TYPE "typeMouldEditor_HMI"
VERSION : 0.1
   STRUCT
      sSelected : Struct   // Selected
         iTool : Int;   // Selected - tool
         sPS : Struct   // Selected - partial shot
            iPS : Int;
            arFlow : Array[0..6] of Real;
            arRatio : Array[0..6] of Real;
            arPressure : Array[0..6] of Real;
            RefComponent : Int;
            "2PoinMovement_Comp01" : Bool;
            "2PoinMovement_Comp02" : Bool;
            "2PoinMovement_Comp03" : Bool;
            "2PoinMovement_Comp04" : Bool;
            "2PoinMovement_Comp05" : Bool;
            "2PoinMovement_Comp06" : Bool;
         END_STRUCT;
         iCalculation : Int;   // Selected - calculation (0=Ftime; 1=flow; 2=weight)
      END_STRUCT;
      arShotSet : Array[0..8] of "UDT925_Shot";   // Shot settings
      uTools : "UDT930_Tool";   // Tool settings
      sCalculatedValues : Struct   // Calculated values
         arTotalFlow : Array[0..8] of Real;   // Calculated values - total flow
      END_STRUCT;
      sStatusBits : Struct   // StatusBits
         xValueChanged : Bool;   // Value changed
         xSafeChanges : Bool;   // Safe changes
         xDiscardChanges : Bool;   // Discard changes
         xDeleteProgram : Bool;   // Delete program
         xFaultDeleteProgram : Bool;   // Fault - delete program
         xProgLoadName : Bool;   // program load name
         xProgLoadNameAckn : Bool;   // program load name - acknowledge
         xFaultValuesnotvalid : Bool;   // values are not valid - flow or shot time wrong
         xPartShotAmount_increase : Bool;   // Partial shot amount - increase
         xPartShotAmount_decrease : Bool;   // Partial shot amount - decrease
      END_STRUCT;
      sColumn : Struct   // Column in HMI
         iShotTime : Int;   // Column - shot time
         iTotalFlow : Int;   // Column - total flow
         iTotalWeight : Int;   // Column - total weight
      END_STRUCT;
      sRow : Struct
         arChangePartialShot : Array[0..8] of Bool;   // Visibility of change partial shot
      END_STRUCT;
   END_STRUCT;
END_TYPE

TYPE "UDT710_EdgeFilter"
TITLE = State of auxiliary drive
VERSION : 0.0
   STRUCT
      Config_Exist : Bool;   // Configuration edge filter existing
      Config_Driven : Bool;   // Configuration with motor
      Config_DifPress : Bool;   // Configuration with difference pressure fault
      Config_Double : Bool;   // Configuration with double egde filter
      RunTime : S5Time;
      PauseTime : S5Time;
      MinTempRelease : Int;   // Min. Temperature to release drive
   END_STRUCT;
END_TYPE

TYPE "UDT100_FeedingPump"
TITLE = State of auxiliary drive
VERSION : 0.0
   STRUCT
      FLT_Exist : Bool;
      FaultLevel_1 : Bool;   // A fault group 1 exist
      FaultLevel_3 : Bool;   // A fault group 3 exist
      Spare0_7 : Bool;
      Reset_Intervall : Bool;   // Reset of intervall- mode at running- and pausetime
      Run : Bool;   // Drive at intervall- mode in running
      Pause : Bool;   // Drive at intervall- mode in pause time
      No_Pausetime : Bool;   // Running- or pausetime is "0" -> drive is running continuously
      Ramp_CVoltage_Off : Bool;   // Flag of delay to switch ON after power lost
      Start_Startupdelay : Bool;   // Information delay time to switch ON after power lost is running
      Disable_Start : Bool;   // Information delay time to switch ON after power lost is running
      Switch_Drive_ON_OFF : Bool;   // Switch auxiliary drive ON-OFF (external signal)
      ManipValuePercent : Int;   // Set value to frequency converter
      State_Drive : Int;   // 1->Drive ON; 2->Fault Drive; 3->Drive requested but not on
   END_STRUCT;
END_TYPE

TYPE "UDT710_FeedingPump"
TITLE = State of auxiliary drive
VERSION : 0.0
   STRUCT
      Config_Exist : Bool;   // Feeding pump exist
      Config_WithFC : Bool;   // Feeding pump with frequency converter
      Config_Without_PresControl : Bool;   // Feeding pump with frequency converter without SetVaue
      Config_With_PresControl : Bool;   // Feeding pump with frequency converter without pressure control
      Config_Bypass : Bool;   // Feeding pump and bypass pump
      Config_Filling : Bool;   // Feeding pump and filling pump
      Config_ManualSwitchON : Bool;   // Feeding pump can be switch on in manal mode
      Config_Spare8 : Bool;
      Config_Spare9 : Bool;
      Config_Spare10 : Bool;
      Config_Spare11 : Bool;
      Config_Spare12 : Bool;
      Config_Spare13 : Bool;
      Config_Spare14 : Bool;
      Config_Spare15 : Bool;
      Config_Spare16 : Bool;
      RunTime : S5Time;   // RunTime feeding pump at bypass
      PauseTime : S5Time;   // PauseTime feeding pump at bypass
      MinTempRelease : Int;   // Min. Temperature to release drive
   END_STRUCT;
END_TYPE

TYPE "UDT927_ShotResult5"
VERSION : 0.1
   STRUCT
      "Date" : Date;
      "Time" : Time_Of_Day;
      StationNo : Byte;
      ProgName : String[20];
      MHNo : Byte := 0;   // Mixinghead number
      PartNo : Int;   // Partnumber of shot at tool
      FoamingTime : Real;   // Foaming Time
      PartWeight : Real;   // Part Weight
      "Name" : Array[1..6] of String[13];
      Mixingratio_SET : Array[1..6] of Real;   // Flow for 8 components
      Mixingratio : Array[1..6] of Real;   // Flow for 8 components
      Flow_SET : Array[1..6] of Real;   // Flow for 8 components
      Flow : Array[1..6] of Real;   // Flow for 8 components
      Pressure_SET : Array[1..6] of Real;   // Pressure for 8 components
      Pressure : Array[1..6] of Real;   // Pressure for 8 components
      Temperature_SET : Array[1..6] of Real;   // Pressure for 8 components
      Temperature : Array[1..6] of Real;   // Pressure for 8 components
   END_STRUCT;
END_TYPE

TYPE "ShotDataToMC"
VERSION : 0.1
   STRUCT
      Data_from_MC : Struct
         Communication : Struct
            Data_read : Bool := FALSE;
            SPARE_00 : Bool := FALSE;
            SPARE_01 : Bool := FALSE;
            SPARE_02 : Bool := FALSE;
            SPARE_03 : Bool := FALSE;
            SPARE_04 : Bool := FALSE;
            SPARE_05 : Bool := FALSE;
            SPARE_06 : Bool := FALSE;
            SPARE_07 : Bool := FALSE;
            SPARE_08 : Bool := FALSE;
            SPARE_09 : Bool := FALSE;
            SPARE_10 : Bool := FALSE;
            SPARE_11 : Bool := FALSE;
            SPARE_12 : Bool := FALSE;
            SPARE_13 : Bool := FALSE;
            SPARE_14 : Bool := FALSE;
         END_STRUCT;
      END_STRUCT;
      Data_to_MC : Struct
         Communication : Struct
            New_Data : Bool := FALSE;
            SPARE_01 : Bool := FALSE;
            SPARE_02 : Bool := FALSE;
            SPARE_03 : Bool := FALSE;
            SPARE_04 : Bool := FALSE;
            SPARE_05 : Bool := FALSE;
            SPARE_06 : Bool := FALSE;
            SPARE_07 : Bool := FALSE;
            SPARE_10 : Bool := FALSE;
            SPARE_11 : Bool := FALSE;
            SPARE_12 : Bool := FALSE;
            SPARE_13 : Bool := FALSE;
            SPARE_14 : Bool := FALSE;
            SPARE_15 : Bool := FALSE;
            SPARE_16 : Bool := FALSE;
            SPARE_17 : Bool := FALSE;
            SPARE_2 : Real;
            SPARE_6 : Int := 0;
         END_STRUCT;
         Act_value : Struct
            MH_No : Byte;   // Actual circulation over mixing head
            Spare : Byte;
            Spare_1 : Int;
            Spare_2 : Real;
            Spare_3 : Real;
            Spare_4 : Real;
            Comp : Array[1..2] of Struct   // Actual values from interface
               Flow : Real;
               Pressure_MH : Real;
               Temperature_MH : Real;
            END_STRUCT;
         END_STRUCT;
         Shot_data : "Shot_data";
      END_STRUCT;
   END_STRUCT;
END_TYPE

TYPE "PB_TecoCS(CW)e_SW-IW"
TITLE = Teco CSe
VERSION : 0.1
// Setpoint- / Actual value telegram for Teco CSe.
// 6word simple protokoll
   STRUCT
      SW : "PB_TecoCS(CW)e_SW";
      IW : "PB_TecoCS(CW)e_IW";
   END_STRUCT;
END_TYPE

TYPE "UDT_State_GWK"
VERSION : 0.1
   STRUCT
      on : Bool;   // Tempering unit is running
      Fault : Bool;   // Fault active
      Weekend_mode : Bool;   // Weekend mode active
      Spare_0_3 : Bool;
      Spare_0_4 : Bool;
      Spare_0_5 : Bool;
      Spare_0_6 : Bool;
      Spare_0_7 : Bool;
      Set_value_tempering_unit : Int;   // Set value for tool temperature
      Act_value_tempering_unit : Real;   // Act value from tempering unit
      Act_value_tool : Int;   // Act value from tool
      Fault_index : Int;   // Index for alarm state
      Fault_state : Word;   // For alarm list
   END_STRUCT;
END_TYPE

TYPE "PB_TecoCS(CW)e_IW"
VERSION : 0.1
   STRUCT
      T1_W1 : Struct   // Telegram 1 word 1 binary encoded
         Bit8 : Bool;   // 1 = Filling level monitoring triggered (M)
         Bit9 : Bool;   // 1 = Pump error motor protection triggered (M)
         Bit10 : Bool;   // 1 = (CS)=Heating error/temperature limiter triggered | (CW)=low pessure switch triggered (M)
         Bit11 : Bool;   // 1 = sensor rupture flow line (M)
         Bit12 : Bool;   // 1 = sensor rupture external sensor (M) (option)
         Bit13 : Bool;   // 1 = Maximum flow line temperature exceeded (P) (only CS)
         Bit14 : Bool;   // 1 = Miniimum flow line temperature exceeded (P)
         Bit15 : Bool;   // Reserve
         Bit0 : Bool;   // 1 = machine operating
         Bit1 : Bool;   // 1 = collective alarm process (P)
         Bit2 : Bool;   // 1 = collective alarm machine (M)
         Bit3 : Bool;   // 1 = error controls/regulator (M)
         Bit4 : Bool;   // 1 = incorrect input setpoint (P)
         Bit5 : Bool;   // 1 = limit violation + (actual value > setpoint + upper limit) (P)
         Bit6 : Bool;   // 1 = limit violation - (actual value < setpoint - lower limit) (P)
         Bit7 : Bool;   // Reserve
      END_STRUCT;
      T1_W2 : Struct   // Telegram 1 word 2 binary encoded
         Bit8 : Bool;   // Reserve
         Bit9 : Bool;   // Reserve
         Bit10 : Bool;   // Reserve
         Bit11 : Bool;   // Reserve
         Bit12 : Bool;   // Reserve
         Bit13 : Bool;   // Reserve
         Bit14 : Bool;   // Reserve
         Bit15 : Bool;   // Reserve
         Bit0 : Bool;   // 1 = interface operation 0 = manual operation
         Bit1 : Bool;   // 1 = External temperature sensor active (option)
         Bit2 : Bool;   // 1 = Machine in normal operation; pump clockwise
         Bit3 : Bool;   // 1 = Standby operation active
         Bit4 : Bool;   // 1 = Machine cools down to switch-off temperature and then switches off
         Bit5 : Bool;   // 1 = Leak stop operation active; pump counter clockwise
         Bit6 : Bool;   // 1 = Mould draining active; pump counter clockwise
         Bit7 : Bool;   // Reserve
      END_STRUCT;
      T1_W3 : Int;   // Temperatur flow line [1/10°C]
      T1_W4 : Int;   // Temperature of the external sensor [1/10°C] (option)
      T1_W5 : Int;   // Flow quantity (option) [1/10 l/m]
      T1_W6 : Int;   // Heating / cooling capacity (option) [1/10%]
   END_STRUCT;
END_TYPE

TYPE "PB_TecoCS(CW)e_SW"
VERSION : 0.1
   STRUCT
      W1 : Struct   // Word 1 binary encoded
         Bit8 : Bool;   // Reserve
         Bit9 : Bool;   // Reserve
         Bit10 : Bool;   // Reserve
         Bit11 : Bool;   // Reserve
         Bit12 : Bool;   // Reserve
         Bit13 : Bool;   // Reserve
         Bit14 : Bool;   // Reserve
         Bit15 : Bool;   // Reserve
         Bit0 : Bool;   // 1 = switch on machine
         Bit1 : Bool;   // 1 = switch on ext. temperature sensor (option)
         Bit2 : Bool;   // 1 = switch on normal operation (heating/cooling & pump clockwise rotation)
         Bit3 : Bool;   // 1 = switch on standby operation (heating/cooling off, pump clockwise rotation)
         Bit4 : Bool;   // 1 = switch on leak stop operation, pump counter-clockwise rotation (option)
         Bit5 : Bool;   // 1 = switch on mould draining, pump counter-clockwise rotation (option)
         Bit6 : Bool;   // 1 = cool down unit and switch off
         Bit7 : Bool;   // 1 = switch on monitoring of limit value
      END_STRUCT;
      T1W2 : Int;   // Setpoint water temperature [1/10°C]
      T1W3 : Int;   // Setpoint limit (relative to setpoint) [1/10°C]
      T1W4 : Int;   // Max. permitted flow line temperature [1/10°C"]
      T1W5 : Int;   // Switch-off temperature (option) [1/10°C]
      T1W6 : Int;   // Reserve
   END_STRUCT;
END_TYPE

TYPE "Shot_data"
VERSION : 0.1
   STRUCT
      MH_No : Byte;   // Mixing head number
      Station_No : Byte;   // Station number
      Shot_No : Int;   // Shot number
      DateTime : Date_And_Time;   // Date and time last shot
      ShotTime_act : Real;   // Shot time last shot
      ShotWeight_act : Real;   // Shot weight last shot
      ShotTime_set : Real;   // Set shot time
      ShotWeight_set : Real;   // Set shot weight
      Spare_1 : Real;
      Spare_2 : Real;
      Comp_act : Array[1..2] of Struct   // Component actual values
         Flow : Real;
         Pressure_MH : Real;
         Temperature_MH : Real;
      END_STRUCT;
      Comp_set : Array[1..2] of Struct   // Component set values
         Flow : Real;
         Pressure_MH : Real;
         Temperature_MH : Real;
      END_STRUCT;
   END_STRUCT;
END_TYPE

TYPE "MC_data"
VERSION : 0.1
   STRUCT
      Tool_temperature : Array[0..16] of Real;
      Reaction_time : Time;
      Closing_time : Time;
      Barcode_1 : String[30];
      Barcode_2 : String[30];
   END_STRUCT;
END_TYPE

TYPE "UDT_RT_Betriebsart"
VERSION : 0.1
   STRUCT
      Gueltig : Bool;   // Es wurde eine gültige Betriebsart angewählt (Hand oder Automatik)
      Hand : Bool;   // Steuerspannung eingeschaltet und Hand angewählt
      Automatik : Bool;   // Steuerspannung eingeschaltet und Automatik angewählt
      Reserve_0_3 : Bool;
      Anfahrwarnung : Bool;   // Eine Anfahrwarnung vor dem Starten des Produktionsbetriebes ist aktiv
      FHM_Anfahrwarnung : Bool;   // Flankenhilfsmerker das die Anfahrwarnung gerade abgelaufen ist
      Lampentest : Bool;   // Steuerspannung eingeschaltet und Lampentest aktiviert
      Steuerspannung_ein : Bool;   // Das Signal "Steuerspannung eingeschaltet" ist länger als 1 Sekunde aktiv
      Flanke_BA_Wechsel : Bool;   // Flankenhilfsmerker für die Betriebsartenumschaltung Hand/ Automatik
      Aktiv : Bool;   // Es wurde eine gültige Betriebsart angewählt und Automatik Stop ist quittiert
      Automatik_Stop_ok : Bool;   // Alle Signale für Automatik- Stop wurden quittiert
      Referenzieren : Bool;   // Einrichten der Anlage für den Produktionnsbetrieb
      Start_Produktion : Bool;   // Die Produktion der Anlage soll gestartet werden (bis Position erreicht)
      Produktion : Bool;   // Der Produktionsbetrieb läuft
      Stop_angefordert : Bool;   // Das Stoppen der Anlage bei erreichen der nächsten Positiuon ist angewählt
      Reserve_1_7 : Bool;
   END_STRUCT;
END_TYPE

TYPE "UDT_RT_Takt"
VERSION : 0.0
   STRUCT
      Vorwarnung_1 : Bool;
      Vorwarnung_2 : Bool;
      Taktzeit_beendet : Bool;
      Taktimpuls : Bool;
      Reserve_0_4 : Bool;
      Reserve_0_5 : Bool;
      Reserve_0_6 : Bool;
      Reserve_0_7 : Bool;
      Reserve_1_0 : Bool;
      Reserve_1_1 : Bool;
      Reserve_1_2 : Bool;
      Reserve_1_3 : Bool;
      Reserve_1_4 : Bool;
      Reserve_1_5 : Bool;
      Reserve_1_6 : Bool;
      Reserve_1_7 : Bool;
   END_STRUCT;
END_TYPE

TYPE "UDT_RT_IPOS"
VERSION : 0.0
   STRUCT
      Ausgaenge_an_IPOS : Struct
         DI_00_Start : Bool;   // Ausgang an Umrichter: Starten des Umrichters (bei Automatik und Referenz)
         DI_01_T_plus : Bool;   // Ausgang an Umrichter: Tippen in positive Richtung
         DI_02_T_minus : Bool;   // Ausgang an Umrichter: Tippen in negative Richtung
         DI_03_Mode_Tipp : Bool;   // Ausgang an Umrichter: Betriebsart Tippen ist angewählt
         DI_04_Mode_Ref : Bool;   // Ausgang an Umrichter: Betriebsart Referenzieren ist angewählt
         DI_05_Mode_Auto : Bool;   // Ausgang an Umrichter: Betriebsart Automatik ist angewählt
         DI_06_Funktion4 : Bool;   // Ausgang an Umrichter:
         DI_07_Funktion5 : Bool;   // Ausgang an Umrichter:
         Reglersperre_Freigabe : Bool;   // Ausgang an Umrichter:
         Freigabe_Schnellstop : Bool;   // Ausgang an Umrichter:
         Freigabe_Halt : Bool;   // Ausgang an Umrichter:
         Halteregelung : Bool;   // Ausgang an Umrichter:
         Integrator_Umschaltung : Bool;   // Ausgang an Umrichter:
         Parametersatz_Umschaltg : Bool;   // Ausgang an Umrichter:
         Reset : Bool;   // Ausgang an Umrichter: Zurückseten der Warnungen
         Reserve0_7 : Bool;   // Ausgang an Umrichter:
         Zielposition : DInt;   // Aktuelle Zielposition (in 1/10 Grad)
         Geschwindigkeit : Word;   // Aktuelle Geschwindigkeit (in 1/100 m/s)
         Positive_Rampe : Word;   // Aktuelle Beschleunigungsrampe (in ms)
         Negative_Rampe : Word;   // Aktuelle Verzögerungsrampe (in ms)
      END_STRUCT;
      Eingaenge_von_IPOS : Struct
         DO_00_Reserve : Bool;   // Eingänge vom Umrichter:
         DO_01_Reserve : Bool;   // Eingänge vom Umrichter:
         DO_02_Reserve : Bool;   // Eingänge vom Umrichter:
         DO_03_Reserve : Bool;   // Eingänge vom Umrichter:
         DO_04_Reserve : Bool;   // Eingänge vom Umrichter:
         DO_05_Reserve : Bool;   // Eingänge vom Umrichter:
         DO_06_Reserve : Bool;   // Eingänge vom Umrichter:
         DO_07_Reserve : Bool;   // Eingänge vom Umrichter:
         Endstufe_freigegeben : Bool;   // Eingänge vom Umrichter:
         Umrichter_betriebsbereit : Bool;   // Eingänge vom Umrichter: Der Umrichter ist betriebsbereit
         Ipos_referenziert : Bool;   // Eingänge vom Umrichter: Der Umrichter ist referenziert
         Ziel_erreicht : Bool;   // Eingänge vom Umrichter: Die vorgegebene Position wurde erreicht
         Bremse_offen : Bool;   // Eingänge vom Umrichter:
         Stoerung_Warnung : Bool;   // Eingänge vom Umrichter:
         Endschalter_rechts_aktiv : Bool;   // Eingänge vom Umrichter:
         Endschalter_links_aktiv : Bool;   // Eingänge vom Umrichter:
         Istposition : DInt;   // Aktuelle Position (in 1/10 Grad)
         PEW_04 : Word;
         PEW_06 : Word;
         PEW_08 : Word;
      END_STRUCT;
      Status : Struct
         Flt_Groupe_Exist : Bool;   // Eine Störung steht an
         Fault_Group1_Exist : Bool;   // Eine Störung der Gruppe 1 steht an
         Fault_Group2_Exist : Bool;   // Eine Störung der Gruppe 2 steht an
         Fault_Group3_Exist : Bool;   // Eine Störung der Gruppe 3 steht an
         Spare_0_4 : Bool;
         Spare_0_5 : Bool;
         Spare_0_6 : Bool;
         FHM_STG_Genauhaltini : Bool;   // Flankenhilfsmerker für die Bildung der Störung des Genauhaltesignales
         HM_Block_ZielPos : Bool;   // Hilfsmerker blockieren "Zielpos erreicht" von IPOS/SEW FU
         BA_Tippen : Bool;   // Es wurde die Betriebsart Tippen Hand (pos/neg) // Auto (pos.) angewählt
         BA_Referenzieren : Bool;   // Es wurde die Betriebsart Referenzieren angewählt
         BA_Takt_Automatik : Bool;   // Es wurde die Betriebsart Takten Automatik (nur positiv ein Segment) angewählt
         BA_Produktion : Bool;   // Es wurde die Betriebsart Produktion bei getakteter Anlage angewählt
         BA_Produktion_Kont : Bool;   // Es wurde die Betriebsart Produktion bei nicht getakteter Anlage angewählt
         BA_gueltig : Bool;   // Es wurde eine gültige Betriebsart bei der Anlage angewählt
         Kettenspannung_noetig : Bool;   // Es ist eine Spannung der Kette im Betrieb notwendig
         FHM_BA_Referenzieren : Bool;   // Flankenmerker für das Starten des Referenzier- Betriebes
         FHM_Referenziert : Bool;   // Flankenmerker für das erreiche der Referenzierungs- Position
         IPOS_referenziert : Bool;   // Der Umrichter wurde Referenziert
         Ziel_ermittelt : Bool;   // Es wurde bereits eine Zielposition für den Umrichter ermittelt
         FHM_Auto_Tip : Bool;   // Flankenhilfsmerker für die Positionierung im automatischem Tipbetrieb
         FHM_Auto_kont : Bool;   // Flankenhilfsmerker für die Positionierung eines kontinuierlichen Betriebes
         Stoppen_erkannt : Bool;   // Das Stoppen des kontinuierlichen Betriebes wurde erkannt
         FHM_Block_ZielPos : Bool;   // Flankenmerker blockieren "Zielpos erreicht" von IPOS/SEW FU
         FHM_STG_Start : Bool;   // Flankenmerker für das Ablöschen des Hilfsmerkers Störung des Genauhaltesignals
         FHM_STG_in_Position : Bool;   // Flankenmerker für das Setzen der Störung des Genauhaltesignals
         Genauhalt_war_verlassen : Bool;   // Merker für die Störungsbildung der Genauhalteposition
         HM_STG_Chk_Genauhalt : Bool;   // Merker zum überprüfen des Genauhaltesignals im kontinuierlichem Betrieb
         HM_Chk_Genauhalt_ok : Bool;   // Hilfsmerker das die Kontrolle des Genauhaltesignals abgeschlossen wurde
         FHM_RT_in_Position : Bool;   // Flankenmerker für die Positionserkennung
         RT_in_Position : Bool;   // Die Anlage ist referenziert und befindet sich in einer definierten Position
         RT_dreht : Bool;   // Der Rundtisch befindet sich in einer automatischen Bewegung
         Aktuelle_Position : Int;   // Wert mit der Aktuellen Position innerhalb des Segmentes (in 1/10 Grad)
         Ziel_Position : DInt;   // Wert für die Berechnung und Weitergabe der Zielposition (in 1/10 Grad)
         Ziel_Geschwindigkeit : Int;   // Wert für die aktuell zu verfahrende Geschwindigkeit (in 1/100 m/s)
         Ziel_Beschleunigung : Int;   // Wert für die aktuell zu verwendende Beschleunigungsrampe (in ms)
         Ziel_Verzoegerung : Int;   // Wert für die aktuell zu verwendende Verzögerungsrampe (in ms)
      END_STRUCT;
   END_STRUCT;
END_TYPE

TYPE "UDT_RT_Station_Nr"
VERSION : 0.1
   STRUCT
      Seg_No_Stat_1 : Int;
      Seg_No_Stat_1_alt : Int;
      Bitmuster_Seg_No_Stat_1 : DWord;
      STG_Nummer_unlogisch : Bool;
      STG_Hardwareabschaltung : Bool;
      STG_Wechsel_in_Pos : Bool;
      STG_Reserve_3 : Bool;
      STG_Reserve_4 : Bool;
      STG_Reserve_5 : Bool;
      STG_Reserve_6 : Bool;
      STG_Reserve_7 : Bool;
      FHM_Nummer_gelesen : Bool;
      FHM_RT_Pos : Bool;
      Reserve9_2 : Bool;
      Reserve9_3 : Bool;
      Reserve9_4 : Bool;
      Reserve9_5 : Bool;
      Reserve9_6 : Bool;
      Reserve9_7 : Bool;
   END_STRUCT;
END_TYPE

TYPE "UDT_RT_Kettenspanner"
VERSION : 0.1
   STRUCT
      Schrittnummer : Byte;
      STG_Entlastung : Bool;
      STG_Druckaufbau : Bool;
      Reserve_12 : Bool;
      Reserve_13 : Bool;
      Reserve_14 : Bool;
      Reserve_15 : Bool;
      V_Entlastung : Bool;
      Kette_gespannt : Bool;
   END_STRUCT;
END_TYPE

TYPE "UDT201_WorkLoadStorage"
TITLE = Signal to tansfer datablocks between work- and loadstorage
VERSION : 0.1
   STRUCT
      Request : Bool;
      Busy : Bool;
      Active : Bool;
      TransferRequest : Bool;
      TransferError : Bool;
      DelayRequest : Bool;
      RequestRuning : Bool;
      Spare07 : Bool;
      TransferStatus : Int;
      TransferStatusSaved : Int;
   END_STRUCT;
END_TYPE

TYPE "Counter"
VERSION : 0.1
   STRUCT
      Anzahl : Int;
      Verbrauch_K1 : Real;   // 1 Kommastelle [kg]
      Verbrauch_K2 : Real;   // 1 Kommastelle [kg]
      Verbrauch_K3 : Real;   // 1 Kommastelle [kg]
      Verbrauch_K4 : Real;   // 1 Kommastelle [kg]
      Verbrauch_K5 : Real;   // 1 Kommastelle [kg]
      Verbrauch_K6 : Real;   // 1 Kommastelle [kg]
      Verbrauch_K7 : Real;   // 1 Kommastelle [kg]
      Verbrauch_K8 : Real;   // 1 Kommastelle [kg]
   END_STRUCT;
END_TYPE

TYPE "Fanuc_Status"
VERSION : 0.0
   STRUCT
      RequestAutomatic : Bool;
      RequestManualMode : Bool;
      AutomaticAccepted : Bool;
      EnableFoamingCycle : Bool;
      StartFoamingCycle : Bool;
      ShotTimesReceived : Bool;
      DataTransmitted : Bool;
      DataInvTransmitted : Bool;
      InterfaceOk : Bool;
      Spare1_1 : Bool;
      Spare1_2 : Bool;
      FLT_detected : Bool;
      EscapingProgram : Bool;
      MovementProg1existing : Bool;
      MovementProg2existing : Bool;
      MovementProg3existing : Bool;
      RobotProgNoMould1 : Int;
      RobotProgNoMould2 : Int;
      RobotProgNoMould3 : Int;
      RobotInProgram : Bool;
      FFdoAction_01_to_Open_MH : Bool;
      doAction_01_to_Open_MH : Bool;
      FMNextPartShot : Bool;   // ramp helpflag for activating new movement program / partshot
      FMRobotNotInAuto : Bool;   // ramp helpflag for resetting the signal "Robot not in Auto"
      RobotNotInAuto : Bool;
      StartBlockedDueToFault : Bool;
      CheckSynchronisation : Bool;
      Spare9_0 : Bool;
      FHMReadyToStart : Bool;
      PUPrgChange : Bool;
      WaitLeaveHome : Bool;
      WaitForHome : Bool;
      FHMSyncIni : Bool;
      CheckHome : Bool;
      CheckMovement : Bool;
      HF_NextMouldEnabled : Bool;   // Helpflag: Conveyor in position where movement to next mould can be enabled
      NextMouldEnabled : Bool;   // movement to next mould can be enabled
      HfAutoStopOk : Bool;   // Helpflag for ramp auto stop ok
      IRB_safe : Bool;   // IRB is in safe position for production without the robot
      Spare10_4 : Bool;
      CleaningProgActive : Bool;   // The robot is working in the cleaning program
      SwitchCleaningON_OFF : Bool;   // Switch cleaning program on/off
      SwitchMaintPosON_OFF : Bool;   // Switch maintenance position on/off
      StateCleaning : Byte;   // 1->Drive ON; 2->Fault Drive; 3->Drive requested but not on
      StateMaintPos : Byte;   // 1->Drive ON; 2->Fault Drive; 3->Drive requested but not on
      MCPlaceNumber : Byte;
      MouldNumber : Byte;
      TimeNumber : Byte;
      OffsetForShotTime : Byte;
      StepNumber : Byte;   // Stepnumber for stepchain of robot interface
      Input : "Fanuc_Input";
      Output : "Fanuc_Output";   // area for output signals (signals received from robot)
      Faults : "Fanuc_Faults";
   END_STRUCT;
END_TYPE

TYPE "UDT254_ServoECylinder"
VERSION : 0.1
   STRUCT
      Signalquellen_E_ZSW1 : Struct   // Signalquellen für Zustandswort E_ZSW1
         E_Einschaltbereit : Bool;   // E_Einschaltbereit
         E_Betriebsbereit : Bool;   // E_Betriebsbereit
         E_Betrieb_freigeben : Bool;   // E_Betrieb_freigeben
         E_Stoerung_wirksam : Bool;   // E_Stoerung_wirksam
         E_Kein_AUS2_wirksam : Bool;   // E_Kein_AUS2_wirksam
         Betriebsbereit_Servo_1 : Bool;   // Servo 1 ist betriebsbereit
         E_Einschaltsperre : Bool;   // E_Einschaltsperre
         E_Warnung_wirksam : Bool;   // E_Warnung_wirksam
         Betriebsbereit_Servo_2 : Bool;   // Servo 2 ist betriebsbereit
         E_Fuehrung_gef_zu_PLC : Bool;   // Führung gefordert zu PLC
         Servo1_Mgrenz_oben : Bool;   // Servo 1 Momentengrenze oben
         E_Vorladung_beendet : Bool;   // E_Vorladung_beendet
         E_Netzschuetz_geschloss : Bool;   // Von Netzschuetz_geschlossen
         Servo1_Mgrenz_unten : Bool;   // Servo 1 Momentengrenze unten
         Servo2_Mgrenz_oben : Bool;   // Servo 2 Momentengrenze oben
         Servo2_Mgrenz_unten : Bool;   // Servo 2 Momentengrenze unten
      END_STRUCT;
      Signalziele_E_STW1 : Struct   // Signalquellen für Steuerwort E_STW1
         Ein : Bool;   // Ein (Vorlade-/Netzschütz ein, Impulsfreigbabe möglich)
         A_Kein_AUS2 : Bool;
         A_Reserviert_0_2 : Bool;   // ------------
         A_Betrieb_freigeben : Bool;   // Betrieb freigeben
         A_Reserviert_0_4 : Bool;   // ------------
         A_Motor_Betrieb_sperren : Bool;   // Motorischer Betrieb sperren
         A_Gen_Betrieb_sperren : Bool;   // Generatorischer Betrieb sperren
         A_Stoerung_quittieren : Bool;   // Störungen quittieren
         A_Reserviert_1_0 : Bool;   // ------------
         A_Reserviert_1_2 : Bool;   // ------------
         A_Fuehrung_durch_PLC : Bool;   // Führung durch PLC
         A_Reserviert_1_3 : Bool;   // ------------
         A_Reserviert_1_4 : Bool;   // ------------
         A_Reserviert_1_5 : Bool;   // ------------
         A_Reserviert_1_6 : Bool;   // ------------
         A_Reserviert_1_7 : Bool;   // ------------
      END_STRUCT;
      Speicher_fuer_Stoerungen : Struct
         Servo1_Mgrenz_unten : Bool;   // Servo 1 Momentengrenze unten erreicht
         Servo1_Mgrenz_oben : Bool;   // Servo 1 Momentengrenze oben erreicht
         Servo2_Mgrenz_unten : Bool;   // Servo 2 Momentengrenze unten erreicht
         Servo2_Mgrenz_oben : Bool;   // Servo 2 Momentengrenze oben erreicht
         Betriebsbereit_Servo_1 : Bool;   // Servo 1 ist nicht betriebsbereit
         Betriebsbereit_Servo_2 : Bool;   // Servo 2 ist nicht betriebsbereit
         Reserviert_0_6 : Bool;   // ------------
         Reserviert_0_7 : Bool;   // ------------
         Reserviert_1_0 : Bool;   // ------------
         Reserviert_1_1 : Bool;   // ------------
         Reserviert_1_2 : Bool;   // ------------
         Reserviert_1_3 : Bool;   // ------------
         Reserviert_1_4 : Bool;   // ------------
         Reserviert_1_5 : Bool;   // ------------
         Reserviert_1_6 : Bool;   // ------------
         Reserviert_1_7 : Bool;   // ------------
      END_STRUCT;
      Momentenueberwachung : Struct
         Istwert_Kolben : Int;   // Momentenwert für Kolben 01
      END_STRUCT;
   END_STRUCT;
END_TYPE

TYPE "UDT312_SafetyDevice"
VERSION : 0.1
   STRUCT
      OpeningSelected : Bool;   // Opening of the safety device is selected
      OpeningEnabled : Bool;   // Opening of the safety device is possible
      EdgeButton : Bool;   // Edge of the button to select opening of the safety device
      HFEdgeButton : Bool;   // Help flag for the edge
      EdgeASReset : Bool;   // Edgo of the reset of Auto Stop from this safety device
      HFEdgeASReset : Bool;   // Help flag for the edge
      Spare0_6 : Bool;
      Spare0_7 : Bool;
      Spare1 : Byte;
   END_STRUCT;
END_TYPE

TYPE "UDT315_ShotadjustS"
TITLE = MH adjustment time for each shot at tool
VERSION : 0.1
   STRUCT
      PS1 : Real;   // Correction value part shot 01
      PS2 : Real;   // Correction value part shot 02
      PS3 : Real;   // Correction value part shot 03
      PS4 : Real;   // Correction value part shot 04
      PS5 : Real;   // Correction value part shot 05
      PS6 : Real;   // Correction value part shot 06
      PS7 : Real := 0.0;   // Correction value part shot 07
      PS8 : Real := 0.0;   // Correction value part shot 08
   END_STRUCT;
END_TYPE

TYPE "UDT316_StateShotAdjust"
VERSION : 0.1
   STRUCT
      CorrFact : Real;
      FoamingTime_ProCan : Real;
      LastShottime : Real;
      SetValueForCorr : Real;
      AdrCorrFact : DWord;
      CorrTimeTest : Real;
      ShotCorrActive : Bool;
      HFShotCorr : Bool;
      ShotCorrTest : Bool;
      Spare03 : Bool;
      Spare04 : Bool;
      Spare05 : Bool;
      Spare06 : Bool;
      Spare07 : Bool;
      SpareByte : Byte;
   END_STRUCT;
END_TYPE

TYPE "UDT502_PV_Tank"
TITLE = Process values of a tank (temp., level, pressure, nucleation)
VERSION : 0.1
   STRUCT
      Temp : "UDT910_ProcessValue";
      Level : "UDT910_ProcessValue";
      Pressure : "UDT910_ProcessValue";
      Nucleation : "UDT910_ProcessValue";
      JacketHeater : "UDT910_ProcessValue";
   END_STRUCT;
END_TYPE

TYPE "UDT504_PV_MH"
TITLE = Process values mixinghead
VERSION : 0.1
   STRUCT
      Pressure_Connection : Array[1..6] of "UDT910_ProcessValue";   // Pressure values at mixinghead conncetions
      Temperature_Connection : Array[1..6] of "UDT910_ProcessValue";   // Temperature values at mixinghead connections
      SteeringPiston : "UDT910_ProcessValue";   // Positon of mixinghead steering piston
      CleaningPiston : "UDT910_ProcessValue";   // Positon of mixinghead cleaning piston
      Inerting : "UDT910_ProcessValue";   // Positon of mixinghead cleaning piston
   END_STRUCT;
END_TYPE

TYPE "UDT506_PV_Machine"
TITLE = Process values machine (shot time)
VERSION : 0.1
   STRUCT
      ShotTime : "UDT910_ProcessValue";   // Refernce number of process value shot time
      Discharge : "UDT910_ProcessValue";   // Refernce number of process value total discharge
      PneumaticFlow : "UDT910_ProcessValue";
   END_STRUCT;
END_TYPE

TYPE "UDT508_PV_Metering"
TITLE = Process values metering (flow, pressure, temp., pp, m. ratio)
VERSION : 0.1
   STRUCT
      Flow : "UDT910_ProcessValue";   // Process value flow rate
      Pressure : "UDT910_ProcessValue";   // Process value pressure
      Temperature : "UDT910_ProcessValue";   // Process value temperature
      Pre_Pressure : "UDT910_ProcessValue";   // Process value pre pressure
      MixingRatio : "UDT910_ProcessValue";   // Process value mixing ratio
   END_STRUCT;
END_TYPE

TYPE "UDT509_PV_Plunger"
TITLE = Process values metering plunger (pressure)
VERSION : 0.1
   STRUCT
      PressurePlunger : "UDT910_ProcessValue";   // Process value pressure Plunger 1
      FlowPlunger : "UDT910_ProcessValue";   // Process value flow plunger 1
      TorquePlunger : "UDT910_ProcessValue";   // Process value torque plunger 1
   END_STRUCT;
END_TYPE

TYPE "UDT700_Machine"
TITLE = Parameter of foaming machine
VERSION : 0.1
   STRUCT
      Int_Runtime_Manual : S5Time;   // Interval run time manual mode
      Int_Pausetime_Manual : S5Time;   // Interval pause time manual mode
      Int_Runtime_Auto : S5Time;   // Interval run time automatic mode
      Int_Pausetime_Auto : S5Time;   // Interval pause time automatic mode
      StrokeCounter_KK : Int;   // Stroke counter of piston machine
      SWU_Intervalltime : S5Time;   // Run time SWU after this there is a switcher to the next SWU
      HP_time_after_shot : S5Time;   // Activate time high pressure after shot
      LP_Valve_switchOFF_Delay : S5Time;   // Switch off delay time of the low pressure valve
      PressureBuildUpTime : S5Time;   // Pressure build up time: Used after start of shot cycle
      StandByTime : S5Time;   // Stand by time: Waiting for next shot request after shot end signal
      CtrlChangeTime1 : S5Time;   // Control change time: Time to adjust flow of squence shot if next MH Nr. is like the previous shot
      CtrlChangeTime2 : S5Time;   // Control change time: Time to adjust flow of squence shot if next MH Nr. is different than the previous shot
      Max_ShotTime : S5Time;   // Time value of maximum shot time
      Min_ShotTime : S5Time;   // Time value of the minum shot time
      Max_WaitTime : S5Time;   // Time value of maximum waiting time after shot request to start foaming
      MH_at_Machine : DWord;   // Which mixinghead works at machine, Bit 0-31 corresponds to Mixinghead 1-32
      Comp_at_Machine : Word;   // Which component works at machine, Bit 0-15 corresponds to component 1-16
      CompPiston_at_Machine : Word;   // Which component is metering as piston, Bit 0-15 corresponds to component 1-16
   END_STRUCT;
END_TYPE

TYPE "UDT701_auxiliaryDrive"
TITLE = Parameter of auxiliary drive
VERSION : 0.1
   STRUCT
      RunTime : S5Time;
      PauseTime : S5Time;
      MinTempRelease : Real;   // Min. Temperature to release drive
   END_STRUCT;
END_TYPE

TYPE "UDT702_Tank"
TITLE = Parameter of tank
VERSION : 0.1
   STRUCT
      "Name" : String[20] := 'Kx';
      FillingTimeControl : S5Time;   // Maximum time to fill the tank
      NoShotFilling : Int;   // Set value of shots to start filling
      TimeToStartFilling : S5Time;   // After this time filling starts again
      PreAgitatingTime : S5Time;   // time to agitate medium before start filling
      Density : Int;   // Density [g/l]
      Color : Byte;   // The color of the daytank
      Existing : Bool;   // These tank is exist
      Deselected : Bool;   // These tank is deselected
      DrainTank : Bool;   // Flag to select draining the tank none min level monitoring
      With_Level : Bool;   // Flag to select kind of filling detection
      With_Level_Monitoring : Bool;   // Flag to select leakage monitoring
      WIth_Loading : Bool;
      With_Heating : Bool;
      With_Vacuum : Bool;
      With_Nucleation : Bool;
      With_Heater_Returnline : Bool;
      With_Drain : Bool;   // Leerfahren
      With_ContainerStation : Bool;
      With_BarelStationAgitator : Bool;
      With_CirculationPump : Bool;   // Tank with circulation pump
      With_CirculationPumpDryRun : Bool;   // Tank with dry run protection for circulation pump
      Spare_34_7 : Bool;
      With_Level_3Liq : Bool;
      With_Level_4Liq : Bool;
      With_Level_Probe : Bool;
      With_Level_SMin : Bool;
      With_Level_SMax : Bool;
      With_Triptray : Bool;
      With_Level_Spare7 : Bool;
      With_Level_Spare8 : Bool;
      With_Filling : Bool;
      With_Filling_Valve : Bool;
      With_Filling_2Valve : Bool;
      With_Filling_ShutDown : Bool;
      With_Filling_Switch : Bool;
      With_Filling_Pump : Bool;   // Filling with a filling pump
      With_Filling_DryRun : Bool;   // Filling with dry run protection
      With_Filling_Pentane : Bool;
      With_Tempering : Bool;
      With_Tempering_TempGeraet : Bool;
      With_Tempering_VKaltwasser : Bool;
      With_Tempering_Heizung : Bool;
      With_Tempering_WTRL : Bool;
      With_Tempering_WTmitFischer : Bool;
      With_Tempering_WTBypass : Bool;
      With_Tempering_WTVL : Bool;
      With_BarelStation : Bool;
      With_BarelStation_Zirkulation : Bool;
      With_BarelStation_PnPump : Bool;
      With_BarelStation_ElPump : Bool;
      With_BarelStation_PnRW : Bool;
      With_BarelStation_ElRW : Bool;
      With_BarelStation_Heating : Bool;
      With_BarelStation_HeatingBottom : Bool;
      With_Agitator : Bool;
      With_Agitator_Converter : Bool;
      With_Agitator_SetValue : Bool;
      With_Agitator_6SetValue : Bool;
      With_Agitator_Spare5 : Bool;
      With_Agitator_Spare6 : Bool;
      With_Agitator_Spare7 : Bool;
      With_Agitator_Spare8 : Bool;
      TankLevel : "UDT702_Tank_Level";
      Agitator : "UDT710_Agitator";
      Agitator_BarelStation : "UDT710_Agitator";
   END_STRUCT;
END_TYPE

TYPE "UDT703_TemperingControl"
TITLE = Parameter of tempering control (2 point)
VERSION : 0.1
   STRUCT
      Dif_Cooling_ON : Real;   // Difference to switch the cooling mode on
      Dif_Cooling_OFF : Real;   // Difference to switch the cooling mode off
      Dif_Heating_ON : Real;   // Difference to switch the heating mode on
      Dif_Heating_OFF : Real;   // Difference to switch the heating mode on
      Max_Temp : Real;   // Max temperature to stop heating (absolute value)
      Min_Temp : Real;   // Min temperature to stop cooling (absolute value)
   END_STRUCT;
END_TYPE

TYPE "UDT704_Mixinghead"
TITLE = Parameter of mixing head
VERSION : 0.1
   STRUCT
      AmountComponent : Byte;   // Amount of components at the mixinghead?
      MachineNumber : Byte;   // Mixinghead at machine number?
      pRrgNumberManual : Byte;   // Start Program number in Manual
      MH_Active : Bool;   // Mixinghead active
      WithCleaningPiston : Bool;   // The mixinghead is equiped with a cleaning piston
      WithNozzleControl : Bool;   // These mixinghead has an nozzle control for more than one mixinghead
      WithLPCirculation : Bool;   // There is a low pressure circulation at the mixinghead
      WithInterface : Bool;   // There is a kind of interface for this mixinghead
      WithInerting : Bool;   // There is a inert system at these mixinghead
      WithHeating : Bool;   // There is a kind of heating at these mixinghead
      WithMHVenting : Bool;   // There is a kind of ventig at these mixinghead
      NozzleLeakageTest : Bool;   // Leakage test for nozzles is active -> close all nozzles and bypasses
      ShotBreak : Bool;   // Shot cycle with this mixinghead is interruptable
      With99program : Bool;   // Mixinghead with 99 manual programs
      Conf_IntWithRobot : Bool;   // Configuration machine with robot
      Conf_IntWithMC : Bool;   // Configuration machine with mould carrier
      Conf_IntWithPlantInerface : Bool;   // Configuration machine with interface to external plant
      Conf_IntWithCoupler : Bool;   // Configuration interface with DP/DP Coupler
      Conf_IntWithProcessValue : Bool;
      Conf_IntWithTag : Bool;
      Conf_MHDigital : Bool;
      Conf_MHControled : Bool;
      Conf_MHFibre : Bool;
      Conf_MHSpray : Bool;
      Conf_MHSpecial : Bool;
      Spare22 : Bool;
      Spare23 : Bool;
      Spare24 : Bool;
      Spare25 : Bool;
      Spare26 : Bool;
      Spare27 : Bool;
      Spare28 : Bool;
      Spare29 : Bool;
      Spare30 : Bool;
      Spare31 : Bool;
      Openingtime : Real;
      Closingtime : Real;
      NozzelCirc : Byte;
      NozzelShot : Byte;
      NozzleRelease : Byte;
      NozzelForcen : Byte;
      DelayTimeNozzlesOff : S5Time;   // Delay time before nozzles and bypasses are switched off after pumps stop
      Delay_UnLockMHafterShot : S5Time;   // Delay unlock mixinghead after shot
      RunTime_MHLock : S5Time;   // Runtime locking mixinghead
      RunTime_MHUnLock : S5Time;   // Runtime unlocking mixinghead
      Cleaning_Piston : "UDT771_CleaningPiston";
      Steering_Piston : "UDT706_SteeringPiston";   // Steering piston
      Corrvalue : Real;   // Correction of runtime steering piston
      Leading_Comp_No : Int;   // Leading component number to calculate mixing ratio
      MH_Connection : Array[1..6] of "UDT1002_MH_Connection";
   END_STRUCT;
END_TYPE

TYPE "UDT702_Tank_Level"
TITLE = Parameter of tank
VERSION : 0.1
   STRUCT
      Max_Level : Real;   // Max filling level: Fault 1 at piston else fault 3
      Start_Level_Filling : Real;
      Stop_Level_Filling : Real;
      Stop_Level_Agitator : Real;   // Beneath this level no agitating
      Min_Level_Warning : Real;
      Min_Level : Real;
   END_STRUCT;
END_TYPE

TYPE "UDT706_SteeringPiston"
TITLE = Parameter of steeringpiston analog control
VERSION : 0.1
   STRUCT
      T_monitoring_open : S5Time;
      T_monitoring_close : S5Time;
   END_STRUCT;
END_TYPE

TYPE "UDT732_FeedPump"
TITLE = Parameter and configuration of feed pump
VERSION : 0.1
   STRUCT
      RunTime : S5Time;
      PauseTime : S5Time;
      Configuration : Byte;
      MinTempRelease : Int;   // Min. Temperature to release drive
   END_STRUCT;
END_TYPE

TYPE "UDT733_CirculationPump"
TITLE = Parameter and configuration of circulation pump
VERSION : 0.1
   STRUCT
      RunTime : S5Time;
      PauseTime : S5Time;
      Configuration : Byte;
      MinTempRelease : Int;   // Min. Temperature to release drive
   END_STRUCT;
END_TYPE

TYPE "UDT734_HeatConverter"
TITLE = Parameter and configuration of heat converter
VERSION : 0.1
   STRUCT
      RunTime : S5Time;
      PauseTime : S5Time;
      Configuration : Byte;
      MinTempRelease : Int;   // Min. Temperature to release drive
   END_STRUCT;
END_TYPE

TYPE "UDT721_Hydraulic"
TITLE = Parameter of mixinghead hydraulik
VERSION : 0.1
   STRUCT
      Hyd_Filter_supervision : S5Time;
      Hyd_P_Startup : S5Time;
      Hyd_P_Supervision : S5Time;
      Hyd_CP_Time : S5Time;
      Hyd_PressureSwitch : S5Time;
      Hyd_SwitchOFFDelay : S5Time;
   END_STRUCT;
END_TYPE

TYPE "UDT753_MeteringPump"
TITLE = Parameter of metering pump
VERSION : 0.1
   STRUCT
      Flow_State : Word;
      RunTimePumpInterval : S5Time;   // Run time for deselected pumps in interval
      PauseTimePumpInterval : S5Time;   // Pause time for deseleted pumps in interval
      Flow_Index : Word;
      DelayPressureFeedP : S5Time;   // Delay of pressure monitoring by using a feed pump
      DelayRunTimeFeedP : S5Time;   // Delay running time feed pump
      MinTempRelease : Real;   // Min. temperature to start the pump
      Pump_Active : Bool;   // Pump active?
      WithFC : Bool;   // Component pump with frecuency converter
      With_2Point : Bool;
      WithFlowControl : Bool;
      WithoutFlowControl : Bool;
      WithFeedPump : Bool;   // Using a feed pump to generate pre pressure
      WithEdgeFilter : Bool;
      PumDeselectionEnable : Bool;   // Pump can deselected
      PumpDeselected : Bool;   // Pump is deselected for maintenance purposes
      PumpDeselectedInterval : Bool;   // Pump is deselected but should run in interval mode
      WithFischerValveHP : Bool;
      WithFischerValveLP : Bool;
      WithHPHeatExchanger : Bool;
      WithLPHeatExchanger : Bool;
      WithExhauseSystem : Bool;
      WithHeating : Bool;
      WithPipeHeating : Bool;
      WithMinTempRelease : Bool;
      WithFlowFactor : Bool;
      With_1Speed : Bool;
      With_2Speed : Bool;
      WithExternalFan : Bool;
      Spare23 : Bool;
      Spare24 : Bool;
      MachineNumber : Byte;   // Mixinghead at machine number?
      "Name" : String[20] := 'Kx';
      TankNo : Int;   // Number of tank which feeds the pump
      AmountOfHeating : Int;   // Amount of heating systems at these component
      Pulse_per_liter : Real;
      MaxFlowLiter : Real := 16.0;   // Max flow [l/min] * 100
      MinFlowPercent : Real := 10.0;   // Min flow in percent of MaxFlow
      MaxFlowPercent : Real := 100.0;   // Max flow in percent of MaxFlow
      FlowThreshold : Real;   // Flow value to switch over pump (Speed; 2-Point)
      FlowFactor : Real;   // Flow value to switch over pump (Speed; 2-Point)
   END_STRUCT;
END_TYPE

TYPE "UDT761_CylinderManager"
TITLE = Parameter of cylinder manager
VERSION : 0.1
   STRUCT
      Preparation_Cylinder : S5Time;   // Within this time piston has to reach start foaming cycle position
      PausePos_Auto : Int;   // Position of cylinder during pausetime in automatic mode (1 = down)
      PausePos_Manual : Int;   // Position of cylinder during pausetime in manual mode (1 = down)
      reserve_01 : Int;
      reserve_02 : Int;
      reserve_03 : Int;
   END_STRUCT;
END_TYPE

TYPE "UDT762_Cylinder"
TITLE = Parameter of metering cylinder
VERSION : 0.1
   STRUCT
      Cyl_PausePosition_Auto : Bool;   // Position of the cylinder during pause in automatic mode (1=below)
      Cyl_PausePosition_Manual : Bool;   // Position of the cylinder during pause in manual mode
      Spare_02 : Bool;
      Spare_03 : Bool;
      Spare_04 : Bool;
      Spare_05 : Bool;
      Spare_06 : Bool;
      Spare_07 : Bool;
      No_cyl_cycle_lubricate : Int;   // Number of cylinder cycle before lubricating
      Spare_6 : Int;
      Spare_8 : Int;
      T_SetValMeterAfterValve : S5Time;   // Time set value metering after valve
      T_ValveMeterAfterSetVal : S5Time;   // Time valve metering after set value
      T_PistonVenting : S5Time;   // Time venting hydraulic between metering and filling
      T_PauseAfterMetering : S5Time;   // Time pause after metering
      T_FillValPreSuctionVal : S5Time;   // Time filling valve before suction valve
      T_SetValFillAfterValve : S5Time;   // Time set value filling after valve
      T_ValveFillAfterSetVal : S5Time;   // Time valve filling after set value
      T_PauseAfterFilling : S5Time;   // Time pause after filling
      T_MonitoringPBFeedpump : S5Time;   // Time monitoring pressure build up feedpump
      Spare26 : Int;
      SetValueFilling : DInt;   // Set value cylinder filling
      SetVMeteringCylSer : DInt;   // Set value cylinder metering during cylinder service
      SetVFillingCylSer : DInt;   // Set value cylinder filling during cylinder service
   END_STRUCT;
END_TYPE

TYPE "UDT771_CleaningPiston"
TITLE = Parameter of mixinghead cleaning piston